// TIA Portal project "proiect" (V17)

(* hardware
DEVICE "S7-1500/ET200MP station_1"  S7-1500 station
   slot 0: "Rail_0"  Rack  6ES7 590-1***0-0AA0
   slot 0: "PS 60W 24/48/60VDC_1"  PS 60W 24/48/60VDC  6ES7 505-0RA00-0AB0  V1.0
   slot 1: "PLC_1"  CPU 1511C-1 PN  6ES7 511-1CK01-0AB0  V2.5
      slot 3: "CPU display_1"  6ES7591-1AA00-0AA0
      slot 32768: "PROFINET interface_1"  X1
         slot 32769: "Port_1"  X1 P1
         slot 32770: "Port_2"  X1 P2
DEVICE "HMI_1"  KTP700 Basic PN
   slot 0: "HMI_1"  KTP700 Basic PN  6AV2 123-2GB03-0AX0  15.1.0.0
   slot 1: "HMI_RT_1"  KTP700 Basic PN  6AV2 123-2GB03-0AX0  15.1.0.0
   slot 5: "HMI_1.IE_CP_1"  PROFINET Interface  15.0.1.0
      slot 1: "PROFINET Interface_1"  PROFINET Interface
         slot 1: "Port_1"  Port
*)

// ===== PLC "PLC_1"  CPU 1511C-1 PN =====

VAR_GLOBAL   // PLC tag table "Default tag table"
   "Tag_1" AT %M10.3 : Bool;
   "Tag_2" AT %M10.4 : Bool;
   "S-R ciuperca" AT %M3.1 : Bool;
   "Tag_4" AT %M3.2 : Bool;
   "Tag_5" AT %M3.3 : Bool;
   "Tag_6" AT %M450.0 : Bool;
   "Tag_7" AT %M450.1 : Bool;
   "Tag_8" AT %M450.2 : Bool;
   "Tag_9" AT %M450.3 : Bool;
   "Tag_10" AT %M450.4 : Bool;
   "Tag_3" AT %M500.0 : Bool;
END_VAR

VAR_GLOBAL   // PLC tag table "Inputs"
   "LS.  mixer_spate" AT %I10.5 : Bool;   // limit switch capat de cursa spate/stanga(mixer)
   "LS. mixer_fata" AT %I10.2 : Bool;   // limit switch capat de cursa fata/dreapta(mixer)
   "LS. loading" AT %I10.7 : Bool;   // limit switch vas pozitionat pe plita
   "LS. unloading" AT %I10.3 : Bool;   // 100% cand versi prod. final
   "LS. mixer_sus" AT %I10.6 : Bool;   // limit switch mixer deasupra bolului de mixare
   "LS. mixer_jos" AT %I10.1 : Bool;   // limit switch mixer in bolul de mixare
END_VAR

VAR_GLOBAL   // PLC tag table "Outputs"
   "ON_OFF plita" AT %Q4.0 : Bool;   // releu plita
   "ON_OFF mixer" AT %Q4.1 : Bool;   // releu mixer
   "ON_OFF pompa_apa" AT %Q4.2 : Bool;   // releu pompa
END_VAR

VAR_GLOBAL   // PLC tag table "Var standard"
   "Clock_Byte" AT %MB0 : Byte;
   "Clock_10Hz" AT %M0.0 : Bool;
   "Clock_5Hz" AT %M0.1 : Bool;
   "Clock_2.5Hz" AT %M0.2 : Bool;
   "Clock_1.25Hz" AT %M0.4 : Bool;
   "Clock_2Hz" AT %M0.3 : Bool;
   "Clock_1Hz" AT %M0.5 : Bool;
   "Clock_0.625Hz" AT %M0.6 : Bool;
   "System_Byte" AT %MB1 : Byte;
   "FirstScan" AT %M1.0 : Bool;
   "Clock_0.5Hz" AT %M0.7 : Bool;
   "DiagStatusUpdate" AT %M1.1 : Bool;
   "AlwaysTRUE" AT %M1.2 : Bool;
   "AlwaysFALSE" AT %M1.3 : Bool;
   "delay1" AT %M200.0 : Bool;
   "delay2" AT %M200.1 : Bool;
   "delay3" AT %M200.2 : Bool;
   "delay4" AT %M200.3 : Bool;
   "delay5" AT %M200.4 : Bool;
   "delay6" AT %M200.5 : Bool;
   "delay7" AT %M200.6 : Bool;
END_VAR

VAR_GLOBAL   // PLC tag table "Markers"
   "ON/OFF_servo1" AT %M1.4 : Bool;
   "ON/OFF_servo2" AT %M1.5 : Bool;
   "ON/OFF_servo3" AT %M2.2 : Bool;
   "Man/Auto" AT %M1.6 : Bool;
   "ON/OFF_Servo1_HMI" AT %MW2 : Word;
   "ON/OFF_servo2_HMI" AT %MW4 : Word;
   "ON/OFF_SERVO3_HMI" AT %MW6 : Word;
   "control_stepper1_HMI" AT %MW8 : Word;
   "control_stepper2_HMI" AT %MW10 : Word;
   "control_stepper3_HMI" AT %MW12 : Word;
   "ON/OFF_SERVO4_HMI" AT %MW14 : Word;
   "ON/OFF_SERVO5_HMI" AT %MW16 : Word;
   "ON/OFF_SERVO6_HMI" AT %MW18 : Word;
   "feedback on/off_mixer" AT %M2.0 : Bool;
   "feedback on/off_pompa" AT %M2.1 : Bool;
   "feedback on/off_plita" AT %M2.3 : Bool;
   "Start_Stop Initializare" AT %M2.4 : Bool;
   "Start/Stop proces" AT %M100.0 : Bool;
   "Feedback On/Off Servo C1" AT %MW24 : Word;
   "Feedback On/Off Servo C2" AT %MW26 : Word;
   "Feedback On/Off Servo L1" AT %MW28 : Word;
   "Feedback On/Off Servo L2" AT %MW30 : Word;
   "Feedback On/Off Servo Z1" AT %MW32 : Word;
   "Feedback On/Off Servo Z2" AT %MW34 : Word;
   "Finalizare_initializare" AT %M100.1 : Bool;
   "Temp_citita" AT %MW36 : Word;
   "MResult_ok" AT %M300.1 : Bool;
   "MResult_not_ok" AT %M300.2 : Bool;
END_VAR

// folder: DB-uri

DATA_BLOCK "DB_Messages"   // DB1
{ S7_Optimized_Access := 'TRUE' }
VERSION : 0.1
   VAR
      B001 : Bool;   // Initializare
      B002 : Word;   // Statia e in modul MANUAL!
      B003 : Word;   // Statia e in modul AUTOMAT!
      B004 : Bool;   // Statia e in modul SEMIAUTOMAT!
      B005 : Word;   // Mixer-ul nu e in pozitia de baza!
      B006 : Word;   // Bolul de amestec nu e in pozitia de baza!
      B007 : Bool;   // Bolul de amestec nu e gol!
      B008 : Word;   // Plita nu este oprita!
      B009 : Word;   // Servo1 pornit
      B010 : Word;   // servo2 pornit
      B011 : Word;   // stepper 1 in functionare
      B012 : Word;   // stepper2 in functionare(vertic)
      B013 : Word;   // stepper3 in functionare (basculare)
      B014 : Bool;
      B015 : Bool;
      B016 : Bool;
      B017 : Bool;
      B018 : Bool;
      B019 : Bool;
      B020 : Bool;
   END_VAR
BEGIN
END_DATA_BLOCK

DATA_BLOCK "DB_Markers"   // DB2
{ S7_Optimized_Access := 'TRUE' }
VERSION : 0.1
   VAR
      Limit_stanga : Bool;   // limita spate mixer
      Limit_dreapta : Bool;   // limita fata mixer
      Limit_mixer_sus : Bool;   // limita mixer sus
      Limit_mixer_jos : Bool;   // limita mixer jos
      limit_loading : Bool;   // limita proces in functionare(loading)
      limit_unloading : Bool;   // limita proces dupa functionare(unloading)
      M_machine_ok : Bool;
      Mixer_pozitie_initiala : Bool;   // Mixer positie de baza(in partea stanga)
      Vas_amestec_poz_init : Bool := 0;   // Vas amestec pozitie de baza(pe plita)
      Vas_amestec_gol : Bool;   // Vas amestec gol
      M_errors : Bool;
      M_Auto : Bool := 0;
      M_Manual : Bool;
      Vas_golit : Bool;   // var folosita in fct pt a goli vasul,dupa instr IF
      "Plita oprita" : Bool;
   END_VAR
BEGIN
END_DATA_BLOCK

DATA_BLOCK "DB_03_Read_Arduino"   // DB3
{ S7_Optimized_Access := 'FALSE' }
VERSION : 0.1
   VAR
      temp_citita : Real;   // temp citita de arduino de senzor
   END_VAR
BEGIN
END_DATA_BLOCK

DATA_BLOCK "DB_HMI"   // DB4
{ S7_Optimized_Access := 'TRUE' }
VERSION : 0.1
   VAR
      "MAN/AUTO" : Bool;
      "Nr-pas_auto" : Int;
      "Selectare Reteta" : Int;
   END_VAR
   VAR RETAIN
      "Bypass-pompa" : Bool;
      bypass_plita : Bool;
      bypass_mixer : Bool;
   END_VAR
   VAR
      "nr. reteta neara" : Int;
      "nr.reteta_lapte" : Int;
      "nr.reteta_alune" : Int;
   END_VAR
BEGIN
END_DATA_BLOCK

DATA_BLOCK "FB_AUTO_DB"   // DB5
{ S7_Optimized_Access := 'TRUE' }
VERSION : 0.1
// stored: InstanceOfName FB_AUTO
"FB_AUTO"
BEGIN
END_DATA_BLOCK

DATA_BLOCK "DB_06_Write_Arduino"   // DB6
{ S7_Optimized_Access := 'FALSE' }
VERSION : 0.1
   VAR
      Servo1 : Bool := 0;
      Servo2 : Bool := 0;
      Servo3 : Bool := 0;
      Servo4 : Bool := 0;
      Servo5 : Bool := 0;
      Servo6 : Bool := 0;
      Stepper1_left : Bool := 0;   // stepper_orizontala(mixer:stanga/dreata)
      Stepper1_right : Bool := 0;   // stepper_orizontala(mixer:stanga/dreata)
      Stepper2_up : Bool := 0;   // stepper_verticala(mixer:sus/jos)
      Stepper2_down : Bool := 0;   // stepper_verticala(mixer:sus/jos)
      Stepper3_loading : Bool := 0;   // stepper _unloading(vrasturnare vas)
      Stepper3_unloading : Bool := 0;
   END_VAR
BEGIN
END_DATA_BLOCK

DATA_BLOCK "DB_HMI_buttons"   // DB7
{ S7_Optimized_Access := 'TRUE' }
VERSION : 0.1
   VAR
      "ON/OFF_plita" : Bool := 0;   // 1-ON/0-OFF
      "ON/OFF_mixer" : Bool := 0;   // 1-ON/0-OFF
      "ON/OFF_pompa" : Bool := 0;   // 1-ON/0-OFF
      Reset : Bool;
      STOP : Bool := 0;   // ciuperca
      Reset_ciuperca : Bool := 0;   // buton care apare dupa ce se activeaza ciuperca(doar pentru a se reseta ciuperca)
      Goleste_vasul : Bool;
      "ON/OFF_servo1" : Bool;
      "ON/OFF_servo2" : Bool;
      "ON/OFF_servo3" : Bool;
      "ON/OFF_servo4" : Bool;
      "ON/OFF_servo5" : Bool;
      "ON/OFF_servo6" : Bool;
      Stepper2_up : Bool := 0;   // buton pentru up la mixer
      Stepper2_down : Bool := 0;   // buton down mixer
      Stepper1_left : Bool := 0;   // buton left mixer
      Stepper1_right : Bool := 0;   // buton right mixer
      Stop_stepper1 : Bool := 0;   // buton stop pentru verticala
      Stop_stepper2 : Bool := 0;   // buton stop pentru orizontala
      Stepper3_loading : Bool;   // buton golire vas
      Stepper3_unloading : Bool;   // buton aducere in pozitie initiala
      Stop_stepper3 : Bool;   // buton stop pentru basculare
      R1_neagra : Bool;
      R2_lapte : Bool;
      R3_cu_alune : Bool;
      Reteta_text_list : Int;
      "Start/Stop_proces_auto" : Bool;
      "Start/Stop_initializare" : Bool;
      Curatare : Bool;
      "Initiere proces" : Bool;
   END_VAR
BEGIN
END_DATA_BLOCK

DATA_BLOCK "DB_Markers_Auto"   // DB8
{ S7_Optimized_Access := 'TRUE' }
VERSION : 0.1
   VAR
      MProcessON : Bool;
      Step2_up : Bool;
      M_Failure : Bool;
      Static_1 : Bool;
      "Dev1:Mixer" : Bool;
      "Dev2:Plita" : Bool := 0;
      "Dev3:Pompa" : Bool;
      "Dev4:Vas_pe_plita" : Bool := 1;
      Curatare : Bool;
      step2_down : Bool;
      step1_left : Bool;
      step1_right : Bool;
      step3_loading : Bool;
      step3_unloading : Bool;
      servo1_auto : Bool;
      servo2_auto : Bool;
      servo3_auto : Bool;
      servo4_auto : Bool;
      servo5_auto : Bool;
      servo6_auto : Bool;
   END_VAR
BEGIN
END_DATA_BLOCK

DATA_BLOCK "DB_MessagesTrigger"   // DB9
{ S7_Optimized_Access := 'TRUE' }
VERSION : 0.1
   VAR
      Info1 : Bool;   // B001:Initializare
      Info2 : Bool;   // B002: Statia e in modul Manual!
      Info3 : Bool;   // B003:Statia e in modul Automat!
      Info4 : Bool;   // B004:Statia e in modul Semiautomat!
      Info5 : Bool;   // B005:Mixerul nu e in pozitia de baza!
      Info6 : Bool;   // B006:Bolul de amestec nu e in pozitia de baza!
      Info7 : Bool;   // B007:Bolul de amestec nu e gol!
      Info8 : Bool;   // B008: Plita nu este oprita!
      Info9 : Bool;
      Info10 : Bool;
      Info11 : Bool;
      Info12 : Bool;
      Info13 : Bool;
      Info14 : Bool;
      Info15 : Bool;
      Info16 : Bool;
      Info17 : Bool;
      Info18 : Bool;
      Info19 : Bool;
      Info20 : Bool;
      Info21 : Bool;
   END_VAR
BEGIN
END_DATA_BLOCK

DATA_BLOCK "DB_Errors"   // DB11
{ S7_Optimized_Access := 'TRUE' }
VERSION : 0.1
   VAR
      Oprire_urgenta : Bool;   // Butonul de urgenta e apasat
      "Eroare1:Vas in aer" : Bool;   // Vasul nu e pe pozitia initiala
      "Eroare2:Mixer" : Bool;   // mixerul nu e in pozitia corespunzatoare(de baza sau de lucru)
      "Eroare3:temp plita" : Bool;   // temp citita >250grade=>eroare la plita =>plita oprita
      "Eroare4:Servo oprite" : Bool;   // daca servo nu sunt oprite=> nu se goleste vasul
      "Eroare5:Limit switch" : Bool;
   END_VAR
BEGIN
END_DATA_BLOCK

// folder: System blocks/Program resources

DATA_BLOCK "counter_reteta-neagra"   // DB10
{ S7_Optimized_Access := 'TRUE' }
AUTHOR : Simatic
FAMILY : IEC
NAME : CNTR
VERSION : 1.0
// stored: InstanceOfName IEC_COUNTER
"IEC_COUNTER"
BEGIN
END_DATA_BLOCK

DATA_BLOCK "ccounter_reteta_lapte"   // DB12
{ S7_Optimized_Access := 'TRUE' }
AUTHOR : Simatic
FAMILY : IEC
NAME : CNTR
VERSION : 1.0
// stored: InstanceOfName IEC_COUNTER
"IEC_COUNTER"
BEGIN
END_DATA_BLOCK

DATA_BLOCK "counter_reteta_alune"   // DB13
{ S7_Optimized_Access := 'TRUE' }
AUTHOR : Simatic
FAMILY : IEC
NAME : CNTR
VERSION : 1.0
// stored: InstanceOfName IEC_COUNTER
"IEC_COUNTER"
BEGIN
END_DATA_BLOCK

// folder: (top level)

ORGANIZATION_BLOCK "Main"   // OB1, LAD, ProgramCycle
TITLE = "Main Program Sweep (Cycle)"
{ S7_Optimized_Access := 'TRUE' }
VERSION : 0.1
   VAR_INPUT
      Initial_Call : Bool;   // Initial call of this OB
      Remanence : Bool;   // =True, if remanent data are available
   END_VAR
   VAR_TEMP   // added for the SCL form of the ladder/FBD networks
      _w1 : Bool;
   END_VAR
BEGIN

REGION Network 1
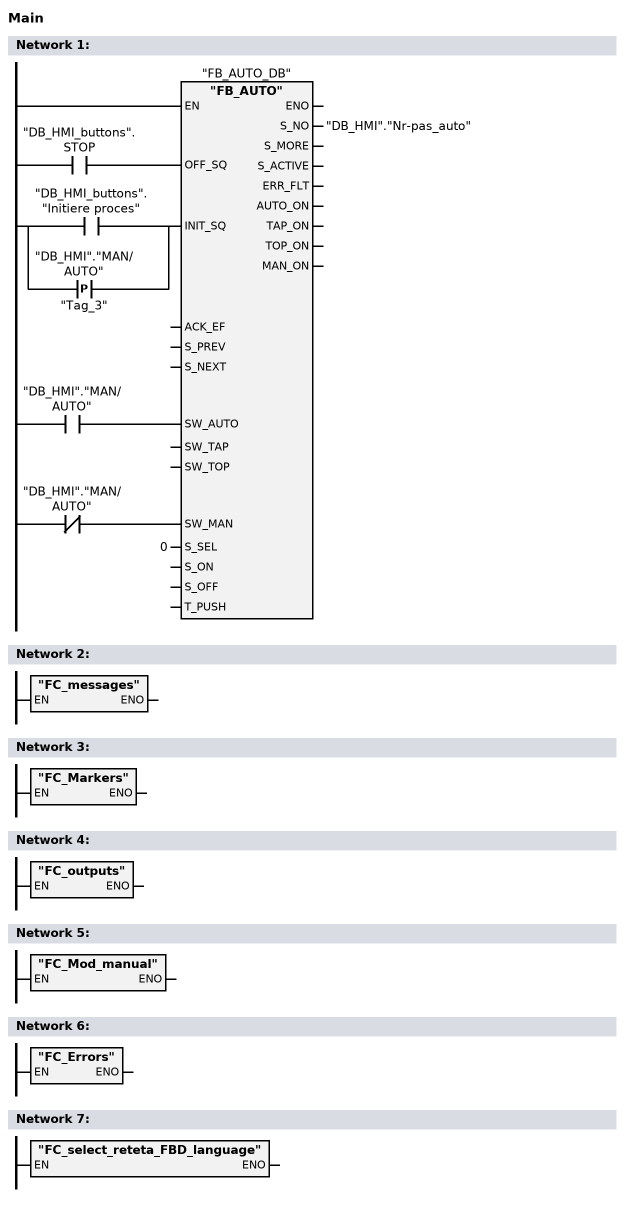
   RUNG wire#powerrail
      "FB_AUTO_DB"(OFF_SQ := wire#w1, INIT_SQ := wire#w2, SW_AUTO := wire#w3, SW_MAN := wire#w4, ACK_EF :=, S_PREV :=, S_NEXT :=, SW_TAP :=, SW_TOP :=, S_SEL := 0, S_ON :=, S_OFF :=, T_PUSH :=, S_NO => "DB_HMI"."Nr-pas_auto", S_MORE =>, S_ACTIVE =>, ERR_FLT =>, AUTO_ON =>, TAP_ON =>, TOP_ON =>, MAN_ON =>)
   END_RUNG
   RUNG wire#powerrail
      Contact( "DB_HMI_buttons".STOP )
   END_RUNG wire#w1
   RUNG wire#powerrail
      Contact( "DB_HMI_buttons"."Initiere proces" )
   END_RUNG wire#w2
   RUNG wire#powerrail
      P_Contact(operand := "DB_HMI"."MAN/AUTO", bit := "Tag_3")
   END_RUNG wire#w2
   RUNG wire#powerrail
      Contact( "DB_HMI"."MAN/AUTO" )
   END_RUNG wire#w3
   RUNG wire#powerrail
      I_Contact( "DB_HMI"."MAN/AUTO" )
   END_RUNG wire#w4
   // the same network as SCL:
   #_w1 := "DB_HMI"."MAN/AUTO" AND NOT "Tag_3";   // rising edge of "DB_HMI"."MAN/AUTO"
   "Tag_3" := "DB_HMI"."MAN/AUTO";
   "FB_AUTO_DB"(OFF_SQ := "DB_HMI_buttons".STOP,   // "FB_AUTO"
                INIT_SQ := "DB_HMI_buttons"."Initiere proces" OR #_w1,
                SW_AUTO := "DB_HMI"."MAN/AUTO",
                SW_MAN := NOT "DB_HMI"."MAN/AUTO",
                S_SEL := 0,
                S_NO => "DB_HMI"."Nr-pas_auto");
END_REGION

REGION Network 2
   RUNG wire#powerrail
      "FC_messages"()
   END_RUNG
   // the same network as SCL:
   "FC_messages"();
END_REGION

REGION Network 3
   RUNG wire#powerrail
      "FC_Markers"()
   END_RUNG
   // the same network as SCL:
   "FC_Markers"();
END_REGION

REGION Network 4
   RUNG wire#powerrail
      "FC_outputs"()
   END_RUNG
   // the same network as SCL:
   "FC_outputs"();
END_REGION

REGION Network 5
   RUNG wire#powerrail
      "FC_Mod_manual"()
   END_RUNG
   // the same network as SCL:
   "FC_Mod_manual"();
END_REGION

REGION Network 6
   RUNG wire#powerrail
      "FC_Errors"()
   END_RUNG
   // the same network as SCL:
   "FC_Errors"();
END_REGION

REGION Network 7
   RUNG wire#powerrail
      "FC_select_reteta_FBD_language"()
   END_RUNG
   // the same network as SCL:
   "FC_select_reteta_FBD_language"();
END_REGION
END_ORGANIZATION_BLOCK

// folder: FB-uri

FUNCTION_BLOCK "FB_AUTO"   // FB1, GRAPH_PLUS
{ S7_Optimized_Access := 'TRUE' }
VERSION : 0.1
   VAR_INPUT
      OFF_SQ : Bool := false;   // Turn sequence off
      INIT_SQ : Bool := false;   // Set sequence to initial state
      ACK_EF : Bool := false;   // Acknowledge all errors and faults
      S_PREV : Bool := false;   // Output previous step in parameter S_NO
      S_NEXT : Bool := false;   // Indicate next step in parameter S_NO
      SW_AUTO : Bool := false;   // Automatic mode
      SW_TAP : Bool := false;   // Semiautomatic/switch with transition
      SW_TOP : Bool := false;   // Semiautomatic/ignore transition
      SW_MAN : Bool := false;   // Manual mode
      S_SEL : Int := 0;   // Select step to be output to S_NO
      S_ON : Bool := false;   // Activate step indicated in S_NO
      S_OFF : Bool := false;   // Deactivate step indicated S_NO
      T_PUSH : Bool := false;   // Enable transition to switch in semi automatic mode
   END_VAR
   VAR_OUTPUT
      S_NO : Int := 0;   // Step number
      S_MORE : Bool := false;   // More steps are available and can be shown in S_NO
      S_ACTIVE : Bool := false;   // Step indicated in S_NO is active
      ERR_FLT : Bool := false;   // Interlock or supervision group error
      AUTO_ON : Bool := false;   // Automatic mode is active
      TAP_ON : Bool := false;   // Semiautomatic mode/step with transition enabled
      TOP_ON : Bool := false;   // Semiautomatic mode/ignore transition enabled
      MAN_ON : Bool := false;   // Manual mode is active
   END_VAR
   VAR
      HMI_INFO : Array[0..9] of UInt;
      IF_PAR : G7_IfParPlus_V6;
      RT_DATA : G7_RTDataPlus_V6;   // Internal data area
      Trans1 : G7_TransitionPlus_V6;   // Transition structure
      Trans2 : G7_TransitionPlus_V6;   // Transition structure
      Trans14 : G7_TransitionPlus_V6;   // Transition structure
      Trans15 : G7_TransitionPlus_V6;   // Transition structure
      Trans16 : G7_TransitionPlus_V6;   // Transition structure
      Trans17 : G7_TransitionPlus_V6;   // Transition structure
      Trans18 : G7_TransitionPlus_V6;   // Transition structure
      Trans19 : G7_TransitionPlus_V6;   // Transition structure
      Trans20 : G7_TransitionPlus_V6;   // Transition structure
      Trans21 : G7_TransitionPlus_V6;   // Transition structure
      Trans22 : G7_TransitionPlus_V6;   // Transition structure
      Trans23 : G7_TransitionPlus_V6;   // Transition structure
      Trans24 : G7_TransitionPlus_V6;   // Transition structure
      Trans25 : G7_TransitionPlus_V6;   // Transition structure
      Trans26 : G7_TransitionPlus_V6;   // Transition structure
      Trans27 : G7_TransitionPlus_V6;   // Transition structure
      Trans28 : G7_TransitionPlus_V6;   // Transition structure
      Trans29 : G7_TransitionPlus_V6;   // Transition structure
      Trans30 : G7_TransitionPlus_V6;   // Transition structure
      Trans35 : G7_TransitionPlus_V6;   // Transition structure
      Trans37 : G7_TransitionPlus_V6;   // Transition structure
      Trans38 : G7_TransitionPlus_V6;   // Transition structure
      Trans39 : G7_TransitionPlus_V6;   // Transition structure
      Trans40 : G7_TransitionPlus_V6;   // Transition structure
      Trans41 : G7_TransitionPlus_V6;   // Transition structure
      Trans42 : G7_TransitionPlus_V6;   // Transition structure
      Trans43 : G7_TransitionPlus_V6;   // Transition structure
      Trans44 : G7_TransitionPlus_V6;   // Transition structure
      Trans45 : G7_TransitionPlus_V6;   // Transition structure
      Trans46 : G7_TransitionPlus_V6;   // Transition structure
      Trans47 : G7_TransitionPlus_V6;   // Transition structure
      Trans48 : G7_TransitionPlus_V6;   // Transition structure
      Trans49 : G7_TransitionPlus_V6;   // Transition structure
      Trans50 : G7_TransitionPlus_V6;   // Transition structure
      Trans51 : G7_TransitionPlus_V6;   // Transition structure
      Trans52 : G7_TransitionPlus_V6;   // Transition structure
      Trans57 : G7_TransitionPlus_V6;   // Transition structure
      Trans58 : G7_TransitionPlus_V6;   // Transition structure
      Trans59 : G7_TransitionPlus_V6;   // Transition structure
      Trans60 : G7_TransitionPlus_V6;   // Transition structure
      Trans64 : G7_TransitionPlus_V6;   // Transition structure
      Trans65 : G7_TransitionPlus_V6;   // Transition structure
      Trans66 : G7_TransitionPlus_V6;   // Transition structure
      Trans67 : G7_TransitionPlus_V6;   // Transition structure
      Trans68 : G7_TransitionPlus_V6;   // Transition structure
      Trans69 : G7_TransitionPlus_V6;   // Transition structure
      Trans70 : G7_TransitionPlus_V6;   // Transition structure
      Trans71 : G7_TransitionPlus_V6;   // Transition structure
      Trans72 : G7_TransitionPlus_V6;   // Transition structure
      Trans73 : G7_TransitionPlus_V6;   // Transition structure
      Trans78 : G7_TransitionPlus_V6;   // Transition structure
      Trans79 : G7_TransitionPlus_V6;   // Transition structure
      Trans80 : G7_TransitionPlus_V6;   // Transition structure
      Trans81 : G7_TransitionPlus_V6;   // Transition structure
      Trans82 : G7_TransitionPlus_V6;   // Transition structure
      Trans83 : G7_TransitionPlus_V6;   // Transition structure
      Trans84 : G7_TransitionPlus_V6;   // Transition structure
      Trans85 : G7_TransitionPlus_V6;   // Transition structure
      Trans86 : G7_TransitionPlus_V6;   // Transition structure
      Trans87 : G7_TransitionPlus_V6;   // Transition structure
      Trans88 : G7_TransitionPlus_V6;   // Transition structure
      Trans89 : G7_TransitionPlus_V6;   // Transition structure
      Trans95 : G7_TransitionPlus_V6;   // Transition structure
      Trans96 : G7_TransitionPlus_V6;   // Transition structure
      Trans98 : G7_TransitionPlus_V6;   // Transition structure
      Trans99 : G7_TransitionPlus_V6;   // Transition structure
      Trans100 : G7_TransitionPlus_V6;   // Transition structure
      Trans101 : G7_TransitionPlus_V6;   // Transition structure
      Trans102 : G7_TransitionPlus_V6;   // Transition structure
      Trans103 : G7_TransitionPlus_V6;   // Transition structure
      Trans104 : G7_TransitionPlus_V6;   // Transition structure
      Trans105 : G7_TransitionPlus_V6;   // Transition structure
      Trans106 : G7_TransitionPlus_V6;   // Transition structure
      Trans107 : G7_TransitionPlus_V6;   // Transition structure
      Trans108 : G7_TransitionPlus_V6;   // Transition structure
      Trans109 : G7_TransitionPlus_V6;   // Transition structure
      Trans112 : G7_TransitionPlus_V6;   // Transition structure
      Trans113 : G7_TransitionPlus_V6;   // Transition structure
      Trans115 : G7_TransitionPlus_V6;   // Transition structure
      Trans116 : G7_TransitionPlus_V6;   // Transition structure
      Trans117 : G7_TransitionPlus_V6;   // Transition structure
      Trans118 : G7_TransitionPlus_V6;   // Transition structure
      Trans119 : G7_TransitionPlus_V6;   // Transition structure
      Trans120 : G7_TransitionPlus_V6;   // Transition structure
      Trans121 : G7_TransitionPlus_V6;   // Transition structure
      Trans122 : G7_TransitionPlus_V6;   // Transition structure
      Trans123 : G7_TransitionPlus_V6;   // Transition structure
      Trans124 : G7_TransitionPlus_V6;   // Transition structure
      Trans125 : G7_TransitionPlus_V6;   // Transition structure
      Trans126 : G7_TransitionPlus_V6;   // Transition structure
      Trans127 : G7_TransitionPlus_V6;   // Transition structure
      Trans128 : G7_TransitionPlus_V6;   // Transition structure
      Trans129 : G7_TransitionPlus_V6;   // Transition structure
      Trans130 : G7_TransitionPlus_V6;   // Transition structure
      Trans134 : G7_TransitionPlus_V6;   // Transition structure
      Trans135 : G7_TransitionPlus_V6;   // Transition structure
      Trans137 : G7_TransitionPlus_V6;   // Transition structure
      Trans138 : G7_TransitionPlus_V6;   // Transition structure
      Trans139 : G7_TransitionPlus_V6;   // Transition structure
      Trans140 : G7_TransitionPlus_V6;   // Transition structure
      Initializare1 : G7_StepPlus_V6;   // Step structure
      "verif poz baza" : G7_StepPlus_V6;   // Step structure
      "on pompa2" : G7_StepPlus_V6;   // Step structure
      Step6 : G7_StepPlus_V6;   // Step structure
      "off pompa+on plita" : G7_StepPlus_V6;   // Step structure
      Step14 : G7_StepPlus_V6;   // Step structure
      Step15 : G7_StepPlus_V6;   // Step structure
      Step16 : G7_StepPlus_V6;   // Step structure
      Step17 : G7_StepPlus_V6;   // Step structure
      Step18 : G7_StepPlus_V6;   // Step structure
      Step19 : G7_StepPlus_V6;   // Step structure
      Step20 : G7_StepPlus_V6;   // Step structure
      Step21 : G7_StepPlus_V6;   // Step structure
      Step22 : G7_StepPlus_V6;   // Step structure
      Step23 : G7_StepPlus_V6;   // Step structure
      Step24 : G7_StepPlus_V6;   // Step structure
      Step25 : G7_StepPlus_V6;   // Step structure
      Step26 : G7_StepPlus_V6;   // Step structure
      Step27 : G7_StepPlus_V6;   // Step structure
      Step28 : G7_StepPlus_V6;   // Step structure
      "Oprire step-poz_init" : G7_StepPlus_V6;   // Step structure
      Step29 : G7_StepPlus_V6;   // Step structure
      Step30 : G7_StepPlus_V6;   // Step structure
      Step34 : G7_StepPlus_V6;   // Step structure
      Step35 : G7_StepPlus_V6;   // Step structure
      Step36 : G7_StepPlus_V6;   // Step structure
      Step37 : G7_StepPlus_V6;   // Step structure
      Step38 : G7_StepPlus_V6;   // Step structure
      Step39 : G7_StepPlus_V6;   // Step structure
      Step40 : G7_StepPlus_V6;   // Step structure
      Step41 : G7_StepPlus_V6;   // Step structure
      Step42 : G7_StepPlus_V6;   // Step structure
      Step43 : G7_StepPlus_V6;   // Step structure
      Step44 : G7_StepPlus_V6;   // Step structure
      Step45 : G7_StepPlus_V6;   // Step structure
      Step46 : G7_StepPlus_V6;   // Step structure
      "Oprire step-poz_init_1" : G7_StepPlus_V6;   // Step structure
      "Activ valve sol prima coloana" : G7_StepPlus_V6;   // Step structure
      delay : G7_StepPlus_V6;   // Step structure
      "off valve" : G7_StepPlus_V6;   // Step structure
      "On plita" : G7_StepPlus_V6;   // Step structure
      timp3 : G7_StepPlus_V6;   // Step structure
      "mixer poz de mixare" : G7_StepPlus_V6;   // Step structure
      "off stepper mix" : G7_StepPlus_V6;   // Step structure
      "On mixer" : G7_StepPlus_V6;   // Step structure
      Step61 : G7_StepPlus_V6;   // Step structure
      "Off mixer" : G7_StepPlus_V6;   // Step structure
      "off plita" : G7_StepPlus_V6;   // Step structure
      "poz initiala mixer" : G7_StepPlus_V6;   // Step structure
      "Oprire step-poz_init_2" : G7_StepPlus_V6;   // Step structure
      "mix-poz_lucru" : G7_StepPlus_V6;   // Step structure
      off_stepper_mix : G7_StepPlus_V6;   // Step structure
      "On mixer2" : G7_StepPlus_V6;   // Step structure
      Step71 : G7_StepPlus_V6;   // Step structure
      "off mixer2" : G7_StepPlus_V6;   // Step structure
      "off plita2" : G7_StepPlus_V6;   // Step structure
      poz_init_MIX : G7_StepPlus_V6;   // Step structure
      "Oprire step-poz_init_3" : G7_StepPlus_V6;   // Step structure
      "Mix-poz_baza" : G7_StepPlus_V6;   // Step structure
      "Oprire stepper" : G7_StepPlus_V6;   // Step structure
      Step89 : G7_StepPlus_V6;   // Step structure
      "Error limit switch" : G7_StepPlus_V6;   // Step structure
      Step91 : G7_StepPlus_V6;   // Step structure
      Step92 : G7_StepPlus_V6;   // Step structure
      Step93 : G7_StepPlus_V6;   // Step structure
      Step90 : G7_StepPlus_V6;   // Step structure
      Step94 : G7_StepPlus_V6;   // Step structure
      Step95 : G7_StepPlus_V6;   // Step structure
      Step96 : G7_StepPlus_V6;   // Step structure
      Step98 : G7_StepPlus_V6;   // Step structure
      Step100 : G7_StepPlus_V6;   // Step structure
      Step101 : G7_StepPlus_V6;   // Step structure
      Step102 : G7_StepPlus_V6;   // Step structure
      Step103 : G7_StepPlus_V6;   // Step structure
      Step104 : G7_StepPlus_V6;   // Step structure
      Step105 : G7_StepPlus_V6;   // Step structure
      Step106 : G7_StepPlus_V6;   // Step structure
      Step107 : G7_StepPlus_V6;   // Step structure
      Step108 : G7_StepPlus_V6;   // Step structure
      Step109 : G7_StepPlus_V6;   // Step structure
      Step110 : G7_StepPlus_V6;   // Step structure
      Step111 : G7_StepPlus_V6;   // Step structure
      Step112 : G7_StepPlus_V6;   // Step structure
      Step113 : G7_StepPlus_V6;   // Step structure
      Step114 : G7_StepPlus_V6;   // Step structure
      Step115 : G7_StepPlus_V6;   // Step structure
      Step116 : G7_StepPlus_V6;   // Step structure
      Step117 : G7_StepPlus_V6;   // Step structure
      Step118 : G7_StepPlus_V6;   // Step structure
      Step121 : G7_StepPlus_V6;   // Step structure
      Step123 : G7_StepPlus_V6;   // Step structure
      Step124 : G7_StepPlus_V6;   // Step structure
      Step125 : G7_StepPlus_V6;   // Step structure
      Step126 : G7_StepPlus_V6;   // Step structure
      SINI : Array[0..2] of USInt;
      LSTT : Array[0..99] of USInt;
      ATAJ : Array[0..99] of USInt;
      ATAB : Array[0..99] of USInt;
      PSTT : Array[0..99] of USInt;
      NSTT : Array[0..99] of USInt;
      ASSJ : Array[0..93] of USInt;
      ASSB : Array[0..93] of USInt;
      PTTS : Array[0..93] of USInt;
      NTTS : Array[0..93] of USInt;
      SW_SQTS : Array[0..93] of USInt;
      SWITCH : Array[0..15] of USInt;
      TVX : Array[0..12] of USInt;
      TTX : Array[0..12] of USInt;
      TSX : Array[0..2] of USInt;
      S00X : Array[0..2] of USInt;
      SOFFX : Array[0..2] of USInt;
      SONX : Array[0..2] of USInt;
      SAX : Array[0..2] of USInt;
      SERRX : Array[0..94] of USInt;
      SMX : Array[0..94] of USInt;
      S0X : Array[0..94] of USInt;
      S1X : Array[0..94] of USInt;
      IL_ALARM_INST : Diag_Alarm;
      SUP_ALARM_INST : Diag_Alarm;
      STEP_TIME_ALARM_INST : Diag_Alarm;
      IEC_TIMER_INST : IEC_TIMER;
      TRANSACTION_FLAG : Bool := false;
   END_VAR
   // SINI[0] := 2;
   // LSTT[0] := 255;
   // LSTT[1] := 255;
   // ATAJ[1] := 1;
   // ATAB[1] := 75;
   // PSTT[1] := 1;
   // NSTT[0] := 1;
   // NSTT[1] := 70;
   // ASSJ[1] := 1;
   // ASSB[1] := 1;
   // PTTS[0] := 255;
   // NTTS[1] := 1;
   // TVX[0] := 16#1;
   // TTX[0] := 16#1;
   // TSX[0] := 16#1;
   // S00X[0] := 16#1;
   // SOFFX[0] := 16#1;
   // SONX[0] := 16#1;
   // SAX[0] := 16#1;
   // SERRX[0] := 16#1;
   // SMX[0] := 16#1;
   // S0X[0] := 16#1;
   // S1X[0] := 16#1;
   // LSTT[2] := 255;
   // LSTT[3] := 255;
   // ATAJ[2] := 2;
   // ATAJ[3] := 3;
   // ATAJ[4] := 4;
   // ATAB[2] := 50;
   // ATAB[3] := 3;
   // ATAB[4] := 4;
   // PSTT[2] := 70;
   // PSTT[3] := 5;
   // PSTT[4] := 6;
   // NSTT[2] := 5;
   // NSTT[3] := 6;
   // ASSJ[2] := 2;
   // ASSJ[3] := 3;
   // ASSJ[4] := 4;
   // ASSB[2] := 2;
   // ASSB[3] := 3;
   // ASSB[4] := 4;
   // PTTS[2] := 50;
   // PTTS[3] := 51;
   // PTTS[4] := 52;
   // NTTS[2] := 51;
   // NTTS[3] := 52;
   // NTTS[4] := 53;
   // LSTT[4] := 255;
   // LSTT[5] := 255;
   // LSTT[6] := 255;
   // LSTT[7] := 255;
   // LSTT[8] := 255;
   // LSTT[9] := 255;
   // LSTT[10] := 255;
   // LSTT[11] := 255;
   // LSTT[12] := 255;
   // LSTT[13] := 255;
   // LSTT[14] := 255;
   // LSTT[15] := 255;
   // LSTT[16] := 255;
   // LSTT[17] := 255;
   // LSTT[18] := 255;
   // LSTT[19] := 255;
   // LSTT[20] := 255;
   // LSTT[21] := 255;
   // LSTT[23] := 255;
   // LSTT[24] := 255;
   // LSTT[25] := 255;
   // LSTT[26] := 255;
   // LSTT[27] := 255;
   // LSTT[28] := 255;
   // LSTT[29] := 255;
   // LSTT[30] := 255;
   // LSTT[31] := 255;
   // LSTT[32] := 255;
   // LSTT[33] := 255;
   // LSTT[34] := 255;
   // LSTT[35] := 255;
   // LSTT[36] := 255;
   // LSTT[37] := 255;
   // LSTT[38] := 255;
   // LSTT[39] := 255;
   // LSTT[40] := 255;
   // LSTT[41] := 255;
   // LSTT[42] := 255;
   // LSTT[44] := 255;
   // LSTT[45] := 255;
   // LSTT[46] := 255;
   // LSTT[47] := 255;
   // LSTT[48] := 255;
   // LSTT[49] := 255;
   // LSTT[50] := 255;
   // LSTT[51] := 255;
   // LSTT[52] := 255;
   // LSTT[53] := 255;
   // LSTT[54] := 255;
   // LSTT[55] := 255;
   // LSTT[56] := 255;
   // LSTT[57] := 255;
   // LSTT[58] := 255;
   // LSTT[59] := 255;
   // LSTT[60] := 255;
   // LSTT[64] := 255;
   // LSTT[62] := 255;
   // LSTT[63] := 255;
   // LSTT[80] := 255;
   // LSTT[66] := 255;
   // LSTT[67] := 255;
   // LSTT[68] := 255;
   // LSTT[69] := 255;
   // LSTT[70] := 255;
   // LSTT[71] := 255;
   // LSTT[72] := 255;
   // LSTT[73] := 255;
   // LSTT[74] := 255;
   // LSTT[75] := 58;
   // LSTT[76] := 255;
   // LSTT[78] := 255;
   // LSTT[79] := 255;
   // LSTT[82] := 255;
   // ATAJ[5] := 5;
   // ATAJ[6] := 6;
   // ATAJ[7] := 7;
   // ATAJ[8] := 8;
   // ATAJ[9] := 9;
   // ATAJ[10] := 10;
   // ATAJ[11] := 11;
   // ATAJ[12] := 12;
   // ATAJ[13] := 13;
   // ATAJ[14] := 14;
   // ATAJ[15] := 15;
   // ATAJ[16] := 16;
   // ATAJ[17] := 17;
   // ATAJ[18] := 18;
   // ATAJ[19] := 19;
   // ATAJ[20] := 20;
   // ATAJ[21] := 21;
   // ATAJ[22] := 22;
   // ATAJ[23] := 23;
   // ATAJ[24] := 24;
   // ATAJ[25] := 25;
   // ATAJ[26] := 26;
   // ATAJ[27] := 27;
   // ATAJ[28] := 28;
   // ATAJ[29] := 29;
   // ATAJ[30] := 30;
   // ATAJ[31] := 31;
   // ATAJ[32] := 32;
   // ATAJ[33] := 33;
   // ATAJ[34] := 34;
   // ATAJ[35] := 35;
   // ATAJ[36] := 36;
   // ATAJ[37] := 37;
   // ATAJ[38] := 38;
   // ATAJ[39] := 39;
   // ATAJ[40] := 40;
   // ATAJ[41] := 41;
   // ATAJ[42] := 42;
   // ATAJ[43] := 43;
   // ATAJ[44] := 44;
   // ATAJ[45] := 45;
   // ATAJ[46] := 46;
   // ATAJ[47] := 47;
   // ATAJ[48] := 48;
   // ATAJ[49] := 49;
   // ATAJ[50] := 50;
   // ATAJ[51] := 51;
   // ATAJ[52] := 52;
   // ATAJ[53] := 53;
   // ATAJ[54] := 54;
   // ATAJ[55] := 55;
   // ATAJ[56] := 56;
   // ATAJ[57] := 57;
   // ATAJ[58] := 58;
   // ATAJ[59] := 59;
   // ATAJ[60] := 60;
   // ATAJ[61] := 61;
   // ATAJ[62] := 62;
   // ATAJ[63] := 63;
   // ATAJ[64] := 64;
   // ATAJ[65] := 65;
   // ATAJ[66] := 66;
   // ATAJ[67] := 67;
   // ATAJ[68] := 68;
   // ATAJ[69] := 69;
   // ATAJ[70] := 70;
   // ATAJ[71] := 71;
   // ATAJ[72] := 72;
   // ATAJ[73] := 73;
   // ATAJ[74] := 74;
   // ATAJ[75] := 75;
   // ATAJ[76] := 76;
   // ATAJ[77] := 77;
   // ATAJ[78] := 78;
   // ATAJ[79] := 79;
   // ATAJ[80] := 80;
   // ATAJ[81] := 81;
   // ATAB[5] := 5;
   // ATAB[6] := 6;
   // ATAB[7] := 7;
   // ATAB[8] := 8;
   // ATAB[9] := 9;
   // ATAB[10] := 10;
   // ATAB[11] := 11;
   // ATAB[12] := 12;
   // ATAB[13] := 13;
   // ATAB[14] := 14;
   // ATAB[15] := 15;
   // ATAB[16] := 16;
   // ATAB[17] := 17;
   // ATAB[18] := 18;
   // ATAB[19] := 2;
   // ATAB[20] := 20;
   // ATAB[21] := 21;
   // ATAB[22] := 22;
   // ATAB[23] := 23;
   // ATAB[24] := 24;
   // ATAB[25] := 25;
   // ATAB[26] := 26;
   // ATAB[27] := 27;
   // ATAB[28] := 28;
   // ATAB[29] := 29;
   // ATAB[30] := 30;
   // ATAB[31] := 31;
   // ATAB[32] := 32;
   // ATAB[33] := 33;
   // ATAB[34] := 34;
   // ATAB[35] := 35;
   // ATAB[36] := 19;
   // ATAB[37] := 37;
   // ATAB[38] := 38;
   // ATAB[39] := 39;
   // ATAB[40] := 40;
   // ATAB[41] := 41;
   // ATAB[42] := 42;
   // ATAB[43] := 43;
   // ATAB[44] := 44;
   // ATAB[45] := 45;
   // ATAB[46] := 46;
   // ATAB[47] := 47;
   // ATAB[48] := 48;
   // ATAB[49] := 49;
   // ATAB[50] := 36;
   // ATAB[51] := 51;
   // ATAB[52] := 52;
   // ATAB[53] := 53;
   // ATAB[54] := 54;
   // ATAB[55] := 55;
   // ATAB[56] := 56;
   // ATAB[57] := 57;
   // ATAB[58] := 58;
   // ATAB[59] := 59;
   // ATAB[60] := 60;
   // ATAB[61] := 61;
   // ATAB[62] := 64;
   // ATAB[63] := 63;
   // ATAB[64] := 62;
   // ATAB[65] := 65;
   // ATAB[66] := 66;
   // ATAB[67] := 67;
   // ATAB[68] := 68;
   // ATAB[69] := 69;
   // ATAB[70] := 70;
   // ATAB[71] := 71;
   // ATAB[72] := 72;
   // ATAB[73] := 73;
   // ATAB[74] := 74;
   // ATAB[75] := 1;
   // ATAB[76] := 76;
   // ATAB[77] := 77;
   // ATAB[78] := 78;
   // ATAB[79] := 79;
   // ATAB[80] := 80;
   // ATAB[81] := 81;
   // PSTT[5] := 7;
   // PSTT[6] := 8;
   // PSTT[7] := 9;
   // PSTT[8] := 10;
   // PSTT[9] := 11;
   // PSTT[10] := 12;
   // PSTT[11] := 13;
   // PSTT[12] := 14;
   // PSTT[13] := 15;
   // PSTT[14] := 16;
   // PSTT[15] := 17;
   // PSTT[16] := 18;
   // PSTT[17] := 19;
   // PSTT[18] := 20;
   // PSTT[19] := 70;
   // PSTT[20] := 21;
   // PSTT[21] := 22;
   // PSTT[22] := 23;
   // PSTT[23] := 24;
   // PSTT[24] := 25;
   // PSTT[25] := 26;
   // PSTT[26] := 27;
   // PSTT[27] := 28;
   // PSTT[28] := 29;
   // PSTT[29] := 30;
   // PSTT[30] := 31;
   // PSTT[31] := 32;
   // PSTT[32] := 33;
   // PSTT[33] := 34;
   // PSTT[34] := 35;
   // PSTT[35] := 36;
   // PSTT[36] := 70;
   // PSTT[37] := 37;
   // PSTT[38] := 38;
   // PSTT[39] := 39;
   // PSTT[40] := 40;
   // PSTT[41] := 41;
   // PSTT[42] := 42;
   // PSTT[43] := 73;
   // PSTT[44] := 44;
   // PSTT[45] := 45;
   // PSTT[46] := 46;
   // PSTT[47] := 47;
   // PSTT[48] := 48;
   // PSTT[49] := 49;
   // PSTT[50] := 70;
   // PSTT[51] := 2;
   // PSTT[52] := 3;
   // PSTT[53] := 4;
   // PSTT[54] := 54;
   // PSTT[55] := 50;
   // PSTT[56] := 51;
   // PSTT[57] := 52;
   // PSTT[58] := 53;
   // PSTT[59] := 55;
   // PSTT[60] := 56;
   // PSTT[61] := 57;
   // PSTT[62] := 58;
   // PSTT[63] := 59;
   // PSTT[64] := 58;
   // PSTT[65] := 61;
   // PSTT[66] := 60;
   // PSTT[67] := 62;
   // PSTT[68] := 63;
   // PSTT[69] := 67;
   // PSTT[70] := 65;
   // PSTT[71] := 66;
   // PSTT[72] := 69;
   // PSTT[73] := 64;
   // PSTT[74] := 68;
   // PSTT[75] := 1;
   // PSTT[76] := 71;
   // PSTT[77] := 72;
   // PSTT[78] := 43;
   // PSTT[79] := 74;
   // PSTT[80] := 75;
   // PSTT[81] := 76;
   // NSTT[4] := 7;
   // NSTT[5] := 8;
   // NSTT[6] := 9;
   // NSTT[7] := 10;
   // NSTT[8] := 64;
   // NSTT[9] := 12;
   // NSTT[10] := 13;
   // NSTT[11] := 14;
   // NSTT[12] := 81;
   // NSTT[13] := 16;
   // NSTT[14] := 17;
   // NSTT[15] := 18;
   // NSTT[16] := 19;
   // NSTT[17] := 20;
   // NSTT[18] := 83;
   // NSTT[19] := 21;
   // NSTT[20] := 22;
   // NSTT[21] := 23;
   // NSTT[23] := 25;
   // NSTT[24] := 26;
   // NSTT[25] := 65;
   // NSTT[26] := 28;
   // NSTT[27] := 29;
   // NSTT[28] := 30;
   // NSTT[29] := 77;
   // NSTT[30] := 32;
   // NSTT[31] := 33;
   // NSTT[32] := 34;
   // NSTT[33] := 35;
   // NSTT[34] := 36;
   // NSTT[35] := 79;
   // NSTT[36] := 37;
   // NSTT[37] := 38;
   // NSTT[38] := 39;
   // NSTT[39] := 60;
   // NSTT[40] := 41;
   // NSTT[41] := 42;
   // NSTT[42] := 43;
   // NSTT[44] := 45;
   // NSTT[45] := 46;
   // NSTT[46] := 47;
   // NSTT[47] := 48;
   // NSTT[48] := 49;
   // NSTT[49] := 75;
   // NSTT[50] := 2;
   // NSTT[51] := 3;
   // NSTT[52] := 4;
   // NSTT[53] := 50;
   // NSTT[54] := 55;
   // NSTT[55] := 51;
   // NSTT[56] := 85;
   // NSTT[57] := 53;
   // NSTT[58] := 54;
   // NSTT[59] := 56;
   // NSTT[60] := 57;
   // NSTT[64] := 61;
   // NSTT[62] := 59;
   // NSTT[63] := 71;
   // NSTT[80] := 76;
   // NSTT[66] := 62;
   // NSTT[67] := 63;
   // NSTT[68] := 40;
   // NSTT[69] := 27;
   // NSTT[70] := 66;
   // NSTT[71] := 67;
   // NSTT[72] := 11;
   // NSTT[73] := 68;
   // NSTT[74] := 69;
   // NSTT[75] := 58;
   // NSTT[76] := 72;
   // NSTT[78] := 73;
   // NSTT[79] := 90;
   // NSTT[82] := 78;
   // ASSJ[5] := 5;
   // ASSJ[6] := 6;
   // ASSJ[7] := 7;
   // ASSJ[8] := 8;
   // ASSJ[9] := 9;
   // ASSJ[10] := 10;
   // ASSJ[11] := 11;
   // ASSJ[12] := 12;
   // ASSJ[13] := 13;
   // ASSJ[14] := 14;
   // ASSJ[15] := 15;
   // ASSJ[16] := 16;
   // ASSJ[17] := 17;
   // ASSJ[18] := 18;
   // ASSJ[19] := 19;
   // ASSJ[20] := 20;
   // ASSJ[21] := 21;
   // ASSJ[22] := 22;
   // ASSJ[23] := 23;
   // ASSJ[24] := 24;
   // ASSJ[25] := 25;
   // ASSJ[26] := 26;
   // ASSJ[27] := 27;
   // ASSJ[28] := 28;
   // ASSJ[29] := 29;
   // ASSJ[30] := 30;
   // ASSJ[31] := 31;
   // ASSJ[32] := 32;
   // ASSJ[33] := 33;
   // ASSJ[34] := 34;
   // ASSJ[35] := 35;
   // ASSJ[36] := 36;
   // ASSJ[37] := 37;
   // ASSJ[38] := 38;
   // ASSJ[39] := 39;
   // ASSJ[40] := 40;
   // ASSJ[41] := 41;
   // ASSJ[42] := 42;
   // ASSJ[43] := 43;
   // ASSJ[44] := 44;
   // ASSJ[45] := 45;
   // ASSJ[46] := 46;
   // ASSJ[47] := 47;
   // ASSJ[48] := 48;
   // ASSJ[49] := 49;
   // ASSJ[50] := 50;
   // ASSJ[51] := 51;
   // ASSJ[52] := 52;
   // ASSJ[53] := 53;
   // ASSJ[54] := 54;
   // ASSJ[55] := 55;
   // ASSJ[56] := 56;
   // ASSJ[57] := 57;
   // ASSJ[58] := 58;
   // ASSJ[59] := 59;
   // ASSJ[60] := 60;
   // ASSJ[61] := 61;
   // ASSJ[62] := 62;
   // ASSJ[63] := 63;
   // ASSJ[64] := 64;
   // ASSJ[65] := 65;
   // ASSJ[66] := 66;
   // ASSJ[67] := 67;
   // ASSJ[68] := 68;
   // ASSJ[69] := 69;
   // ASSJ[70] := 70;
   // ASSJ[71] := 71;
   // ASSJ[72] := 72;
   // ASSJ[73] := 73;
   // ASSJ[74] := 74;
   // ASSJ[75] := 75;
   // ASSJ[76] := 76;
   // ASSJ[77] := 77;
   // ASSB[5] := 5;
   // ASSB[6] := 6;
   // ASSB[7] := 7;
   // ASSB[8] := 8;
   // ASSB[9] := 9;
   // ASSB[10] := 10;
   // ASSB[11] := 11;
   // ASSB[12] := 12;
   // ASSB[13] := 13;
   // ASSB[14] := 14;
   // ASSB[15] := 15;
   // ASSB[16] := 16;
   // ASSB[17] := 17;